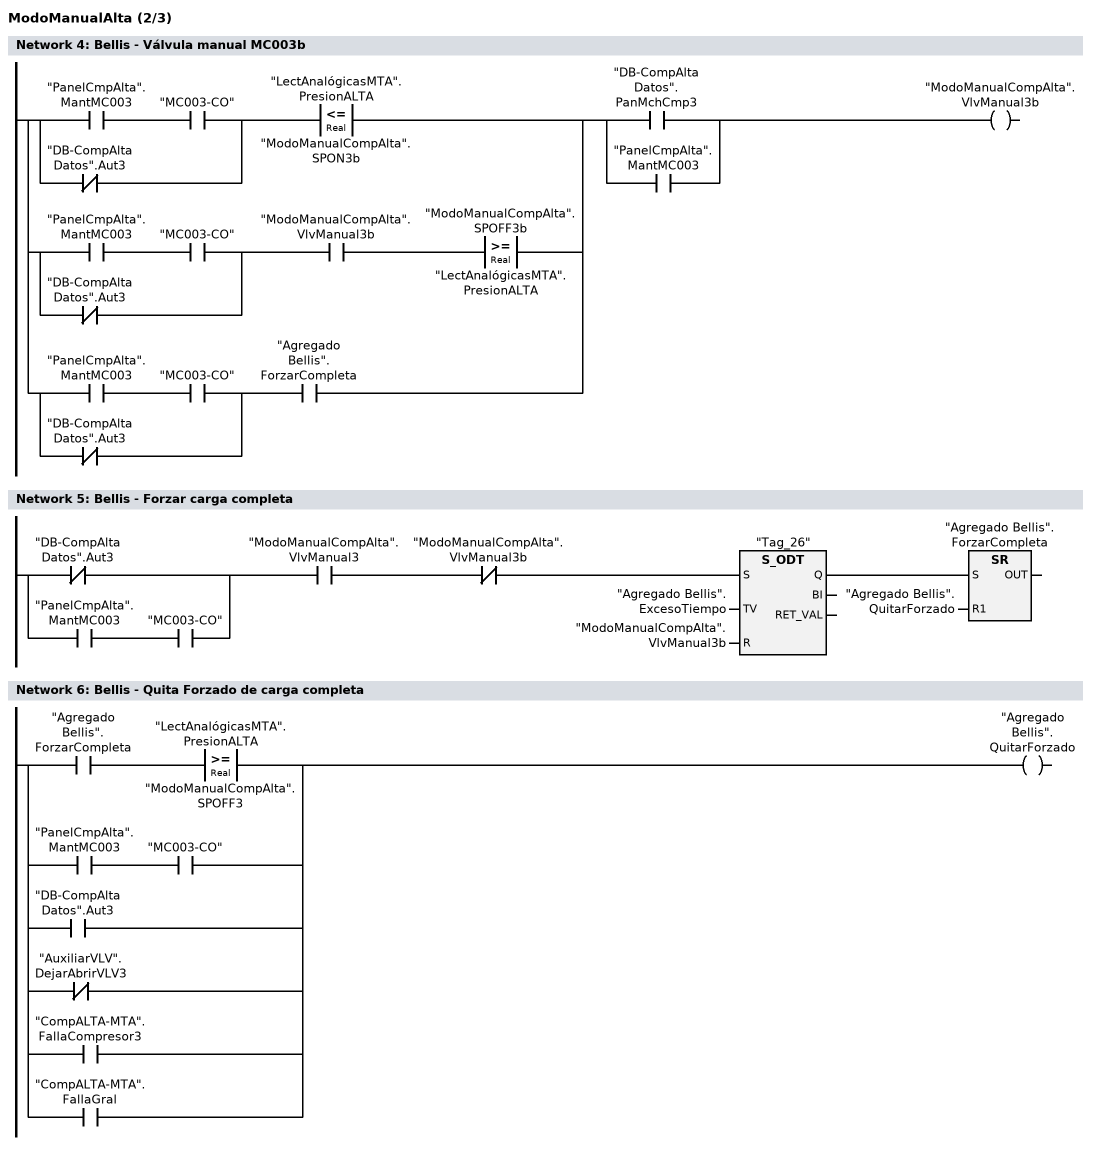
   "ModoManualCompAlta".VlvManual3b := (((NOT "DB-CompAltaDatos".Aut3 OR ("PanelCmpAlta".MantMC003 AND "MC003-CO")) AND ("LectAnalógicasMTA".PresionALTA <= "ModoManualCompAlta".SPON3b)) OR ((NOT "DB-CompAltaDatos".Aut3 OR ("PanelCmpAlta".MantMC003 AND "MC003-CO")) AND "ModoManualCompAlta".VlvManual3b AND ("ModoManualCompAlta".SPOFF3b >= "LectAnalógicasMTA".PresionALTA)) OR ((NOT "DB-CompAltaDatos".Aut3 OR ("PanelCmpAlta".MantMC003 AND "MC003-CO")) AND "Agregado Bellis".ForzarCompleta)) AND ("DB-CompAltaDatos".PanMchCmp3 OR "PanelCmpAlta".MantMC003);
END_REGION

REGION Network 5: Bellis - Forzar carga completa
   RUNG wire#powerrail
      I_Contact( "DB-CompAltaDatos".Aut3 )
      wire#w1
      Contact( "ModoManualCompAlta".VlvManual3 )
      I_Contact( "ModoManualCompAlta".VlvManual3b )
      S_ODT(T_NO := "Tag_26", TV := "Agregado Bellis".ExcesoTiempo, R := "ModoManualCompAlta".VlvManual3b, BI =>, RET_VAL =>)
      S_SR(operand := "Agregado Bellis".ForzarCompleta, r1 := "Agregado Bellis".QuitarForzado)
   END_RUNG
   RUNG wire#powerrail
      Contact( "PanelCmpAlta".MantMC003 )
      Contact( "MC003-CO" )
   END_RUNG wire#w1
   // the same network as SCL:
   #_s5time1 := S_ODT(T_NO := "Tag_26",
                      S := (NOT "DB-CompAltaDatos".Aut3 OR ("PanelCmpAlta".MantMC003 AND "MC003-CO")) AND "ModoManualCompAlta".VlvManual3 AND NOT "ModoManualCompAlta".VlvManual3b,
                      TV := "Agregado Bellis".ExcesoTiempo,
                      R := "ModoManualCompAlta".VlvManual3b,
                      Q => #_w1);
   IF #_w1 THEN
       "Agregado Bellis".ForzarCompleta := TRUE;   // SR flip-flop
   END_IF;
   IF "Agregado Bellis".QuitarForzado THEN "Agregado Bellis".ForzarCompleta := FALSE; END_IF;
END_REGION

REGION Network 6: Bellis - Quita Forzado de carga completa
   "Agregado Bellis".QuitarForzado := ("Agregado Bellis".ForzarCompleta AND ("LectAnalógicasMTA".PresionALTA >= "ModoManualCompAlta".SPOFF3)) OR "DB-CompAltaDatos".Aut3 OR ("PanelCmpAlta".MantMC003 AND "MC003-CO") OR NOT "AuxiliarVLV".DejarAbrirVLV3 OR "CompALTA-MTA".FallaCompresor3 OR "CompALTA-MTA".FallaGral;
END_REGION

REGION Network 7
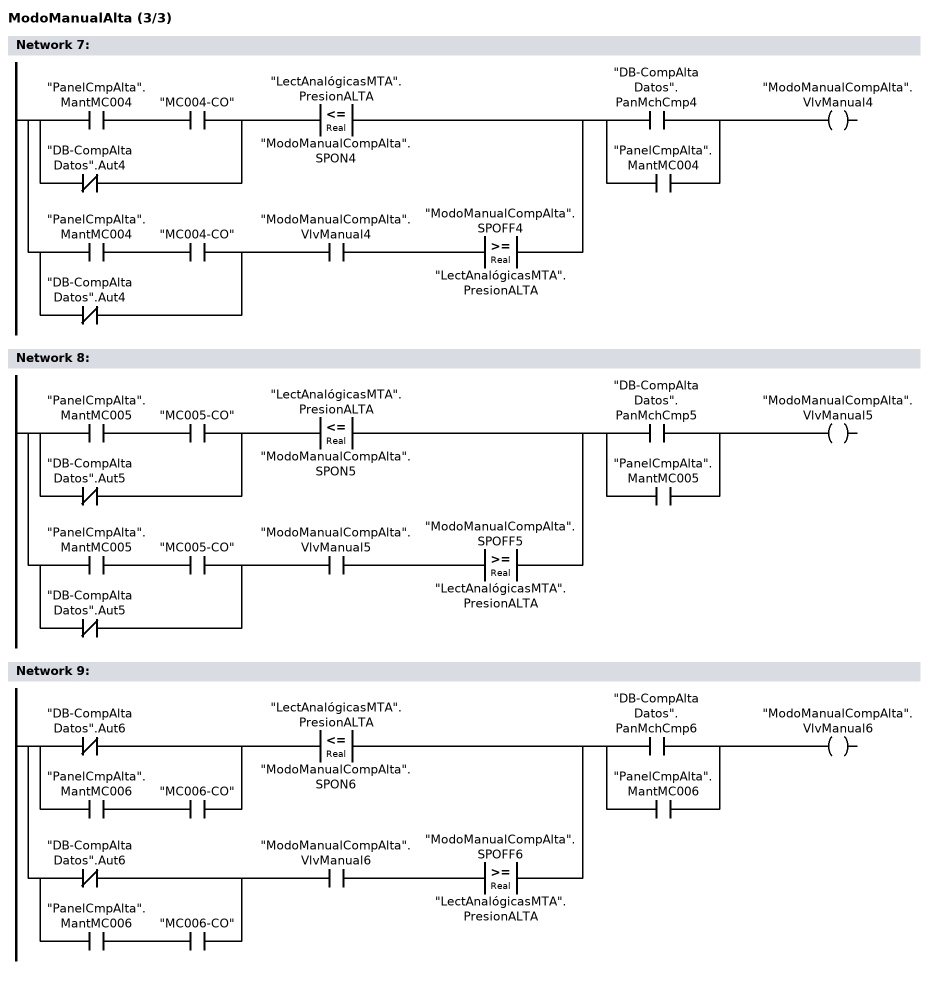
   "ModoManualCompAlta".VlvManual4 := (((NOT "DB-CompAltaDatos".Aut4 OR ("PanelCmpAlta".MantMC004 AND "MC004-CO")) AND ("LectAnalógicasMTA".PresionALTA <= "ModoManualCompAlta".SPON4)) OR ((NOT "DB-CompAltaDatos".Aut4 OR ("PanelCmpAlta".MantMC004 AND "MC004-CO")) AND "ModoManualCompAlta".VlvManual4 AND ("ModoManualCompAlta".SPOFF4 >= "LectAnalógicasMTA".PresionALTA))) AND ("DB-CompAltaDatos".PanMchCmp4 OR "PanelCmpAlta".MantMC004);
END_REGION

REGION Network 8
   "ModoManualCompAlta".VlvManual5 := (((NOT "DB-CompAltaDatos".Aut5 OR ("PanelCmpAlta".MantMC005 AND "MC005-CO")) AND ("LectAnalógicasMTA".PresionALTA <= "ModoManualCompAlta".SPON5)) OR ((NOT "DB-CompAltaDatos".Aut5 OR ("PanelCmpAlta".MantMC005 AND "MC005-CO")) AND "ModoManualCompAlta".VlvManual5 AND ("ModoManualCompAlta".SPOFF5 >= "LectAnalógicasMTA".PresionALTA))) AND ("DB-CompAltaDatos".PanMchCmp5 OR "PanelCmpAlta".MantMC005);
END_REGION

REGION Network 9
   RUNG wire#powerrail
      I_Contact( "DB-CompAltaDatos".Aut6 )
      wire#w1
      { S7_Templates := "SrcType := Real" } LE_Contact(in1 := "LectAnalógicasMTA".PresionALTA, in2 := "ModoManualCompAlta".SPON6)
      wire#w2
      Contact( "DB-CompAltaDatos".PanMchCmp6 )
      wire#w4
      Coil( "ModoManualCompAlta".VlvManual6 )
   END_RUNG
   RUNG wire#powerrail
      Contact( "PanelCmpAlta".MantMC006 )
      Contact( "MC006-CO" )
   END_RUNG wire#w1
   RUNG wire#powerrail
      I_Contact( "DB-CompAltaDatos".Aut6 )
      wire#w3
      Contact( "ModoManualCompAlta".VlvManual6 )
      { S7_Templates := "SrcType := Real" } GE_Contact(in1 := "ModoManualCompAlta".SPOFF6, in2 := "LectAnalógicasMTA".PresionALTA)
   END_RUNG wire#w2
   RUNG wire#powerrail
      Contact( "PanelCmpAlta".MantMC006 )
      Contact( "MC006-CO" )
   END_RUNG wire#w3
   RUNG wire#w2
      Contact( "PanelCmpAlta".MantMC006 )
   END_RUNG wire#w4
   // the same network as SCL:
   "ModoManualCompAlta".VlvManual6 := (((NOT "DB-CompAltaDatos".Aut6 OR ("PanelCmpAlta".MantMC006 AND "MC006-CO")) AND ("LectAnalógicasMTA".PresionALTA <= "ModoManualCompAlta".SPON6)) OR ((NOT "DB-CompAltaDatos".Aut6 OR ("PanelCmpAlta".MantMC006 AND "MC006-CO")) AND "ModoManualCompAlta".VlvManual6 AND ("ModoManualCompAlta".SPOFF6 >= "LectAnalógicasMTA".PresionALTA))) AND ("DB-CompAltaDatos".PanMchCmp6 OR "PanelCmpAlta".MantMC006);
END_REGION
END_FUNCTION

// folder: Compresores/Alta/Máquina de Estados

FUNCTION "LogMaqEstGeneral" : Void   // FC35, LAD
{ S7_Optimized_Access := 'FALSE' }
VERSION : 0.1
BEGIN

REGION Network 1
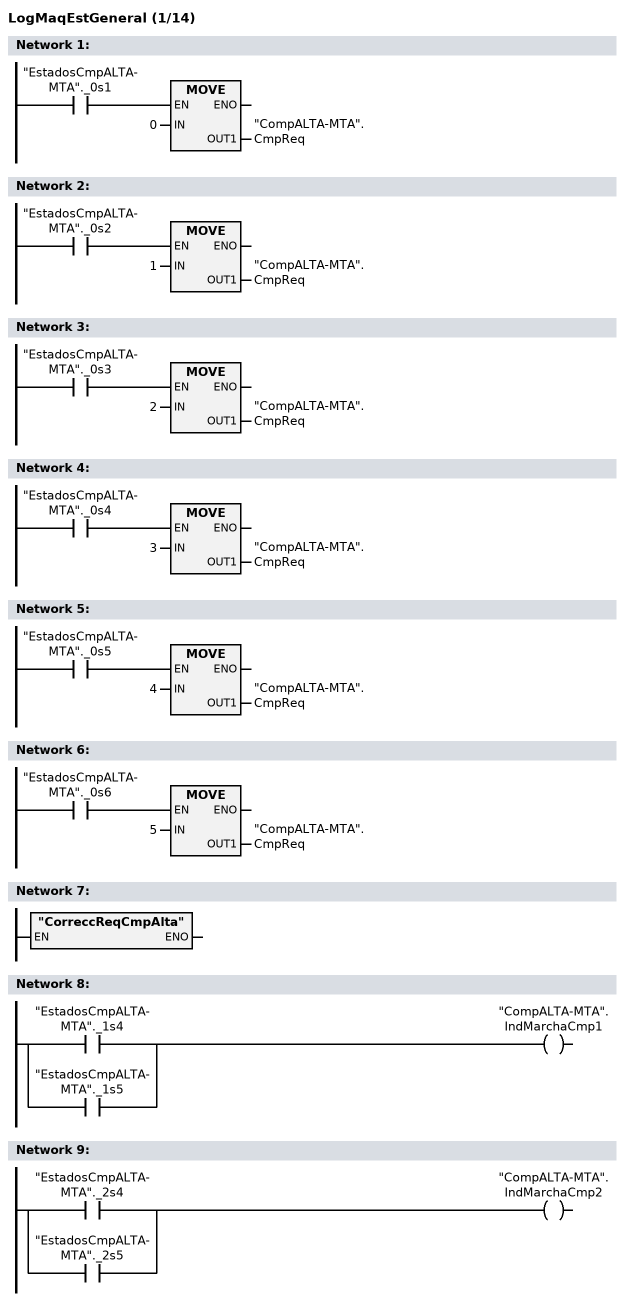
   RUNG wire#powerrail
      Contact( "EstadosCmpALTA-MTA"._0s1 )
      { S7_GenerateENO := "TRUE" } Move(in := 0, out1 => "CompALTA-MTA".CmpReq)
   END_RUNG
   // the same network as SCL:
   IF "EstadosCmpALTA-MTA"._0s1 THEN "CompALTA-MTA".CmpReq := 0; END_IF;
END_REGION

REGION Network 2
   RUNG wire#powerrail
      Contact( "EstadosCmpALTA-MTA"._0s2 )
      { S7_GenerateENO := "TRUE" } Move(in := 1, out1 => "CompALTA-MTA".CmpReq)
   END_RUNG
   // the same network as SCL:
   IF "EstadosCmpALTA-MTA"._0s2 THEN "CompALTA-MTA".CmpReq := 1; END_IF;
END_REGION

REGION Network 3
   RUNG wire#powerrail
      Contact( "EstadosCmpALTA-MTA"._0s3 )
      { S7_GenerateENO := "TRUE" } Move(in := 2, out1 => "CompALTA-MTA".CmpReq)
   END_RUNG
   // the same network as SCL:
   IF "EstadosCmpALTA-MTA"._0s3 THEN "CompALTA-MTA".CmpReq := 2; END_IF;
END_REGION

REGION Network 4
   RUNG wire#powerrail
      Contact( "EstadosCmpALTA-MTA"._0s4 )
      { S7_GenerateENO := "TRUE" } Move(in := 3, out1 => "CompALTA-MTA".CmpReq)
   END_RUNG
   // the same network as SCL:
   IF "EstadosCmpALTA-MTA"._0s4 THEN "CompALTA-MTA".CmpReq := 3; END_IF;
END_REGION

REGION Network 5
   RUNG wire#powerrail
      Contact( "EstadosCmpALTA-MTA"._0s5 )
      { S7_GenerateENO := "TRUE" } Move(in := 4, out1 => "CompALTA-MTA".CmpReq)
   END_RUNG
   // the same network as SCL:
   IF "EstadosCmpALTA-MTA"._0s5 THEN "CompALTA-MTA".CmpReq := 4; END_IF;
END_REGION

REGION Network 6
   RUNG wire#powerrail
      Contact( "EstadosCmpALTA-MTA"._0s6 )
      { S7_GenerateENO := "TRUE" } Move(in := 5, out1 => "CompALTA-MTA".CmpReq)
   END_RUNG
   // the same network as SCL:
   IF "EstadosCmpALTA-MTA"._0s6 THEN "CompALTA-MTA".CmpReq := 5; END_IF;
END_REGION

REGION Network 7
   RUNG wire#powerrail
      "CorreccReqCmpAlta"()
   END_RUNG
   // the same network as SCL:
   "CorreccReqCmpAlta"();
END_REGION

REGION Network 8
   RUNG wire#powerrail
      Contact( "EstadosCmpALTA-MTA"._1s4 )
      wire#w1
      Coil( "CompALTA-MTA".IndMarchaCmp1 )
   END_RUNG
   RUNG wire#powerrail
      Contact( "EstadosCmpALTA-MTA"._1s5 )
   END_RUNG wire#w1
   // the same network as SCL:
   "CompALTA-MTA".IndMarchaCmp1 := "EstadosCmpALTA-MTA"._1s4 OR "EstadosCmpALTA-MTA"._1s5;
END_REGION

REGION Network 9
   RUNG wire#powerrail
      Contact( "EstadosCmpALTA-MTA"._2s4 )
      wire#w1
      Coil( "CompALTA-MTA".IndMarchaCmp2 )
   END_RUNG
   RUNG wire#powerrail
      Contact( "EstadosCmpALTA-MTA"._2s5 )
   END_RUNG wire#w1
   // the same network as SCL:
   "CompALTA-MTA".IndMarchaCmp2 := "EstadosCmpALTA-MTA"._2s4 OR "EstadosCmpALTA-MTA"._2s5;
END_REGION

REGION Network 10
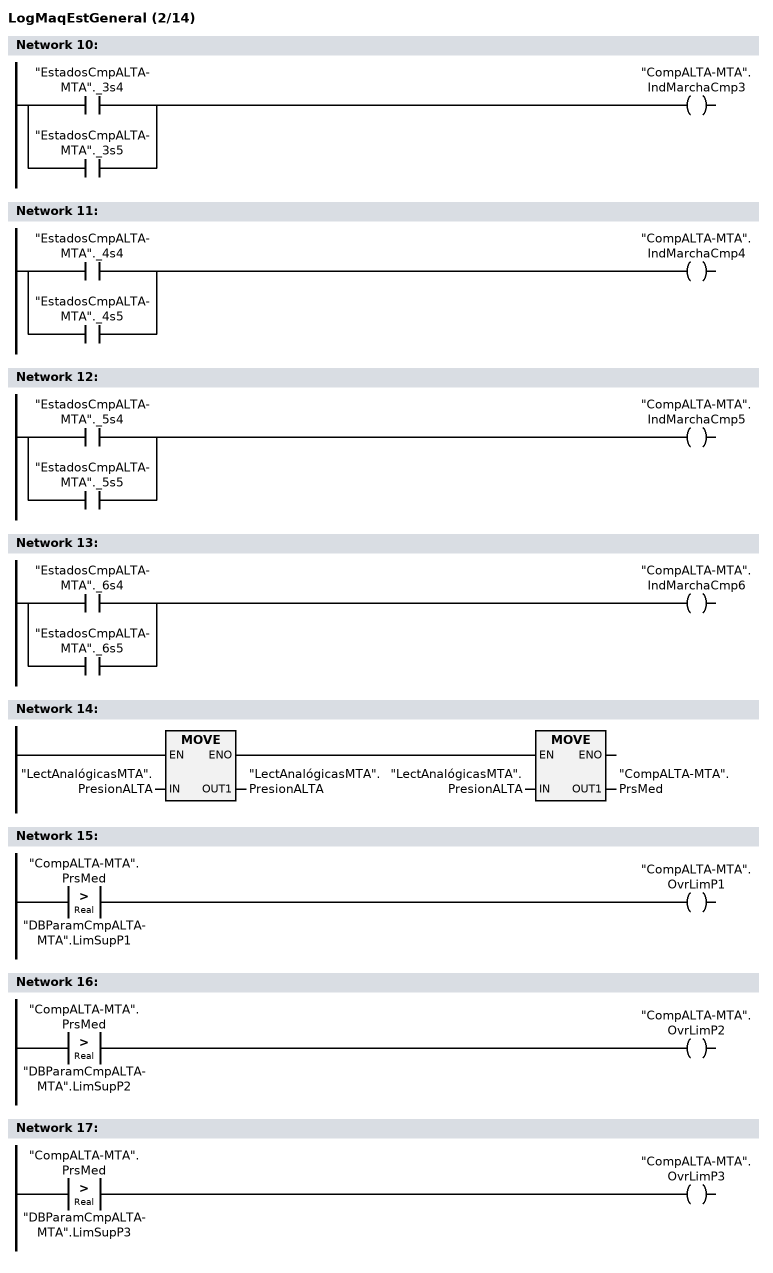
   RUNG wire#powerrail
      Contact( "EstadosCmpALTA-MTA"._3s4 )
      wire#w1
      Coil( "CompALTA-MTA".IndMarchaCmp3 )
   END_RUNG
   RUNG wire#powerrail
      Contact( "EstadosCmpALTA-MTA"._3s5 )
   END_RUNG wire#w1
   // the same network as SCL:
   "CompALTA-MTA".IndMarchaCmp3 := "EstadosCmpALTA-MTA"._3s4 OR "EstadosCmpALTA-MTA"._3s5;
END_REGION

REGION Network 11
   RUNG wire#powerrail
      Contact( "EstadosCmpALTA-MTA"._4s4 )
      wire#w1
      Coil( "CompALTA-MTA".IndMarchaCmp4 )
   END_RUNG
   RUNG wire#powerrail
      Contact( "EstadosCmpALTA-MTA"._4s5 )
   END_RUNG wire#w1
   // the same network as SCL:
   "CompALTA-MTA".IndMarchaCmp4 := "EstadosCmpALTA-MTA"._4s4 OR "EstadosCmpALTA-MTA"._4s5;
END_REGION

REGION Network 12
   RUNG wire#powerrail
      Contact( "EstadosCmpALTA-MTA"._5s4 )
      wire#w1
      Coil( "CompALTA-MTA".IndMarchaCmp5 )
   END_RUNG
   RUNG wire#powerrail
      Contact( "EstadosCmpALTA-MTA"._5s5 )
   END_RUNG wire#w1
   // the same network as SCL:
   "CompALTA-MTA".IndMarchaCmp5 := "EstadosCmpALTA-MTA"._5s4 OR "EstadosCmpALTA-MTA"._5s5;
END_REGION

REGION Network 13
   RUNG wire#powerrail
      Contact( "EstadosCmpALTA-MTA"._6s4 )
      wire#w1
      Coil( "CompALTA-MTA".IndMarchaCmp6 )
   END_RUNG
   RUNG wire#powerrail
      Contact( "EstadosCmpALTA-MTA"._6s5 )
   END_RUNG wire#w1
   // the same network as SCL:
   "CompALTA-MTA".IndMarchaCmp6 := "EstadosCmpALTA-MTA"._6s4 OR "EstadosCmpALTA-MTA"._6s5;
END_REGION

REGION Network 14
   RUNG wire#powerrail
      { S7_GenerateENO := "TRUE" } Move(in := "LectAnalógicasMTA".PresionALTA, out1 => "LectAnalógicasMTA".PresionALTA)
      { S7_GenerateENO := "TRUE" } Move(in := "LectAnalógicasMTA".PresionALTA, out1 => "CompALTA-MTA".PrsMed)
   END_RUNG
   // the same network as SCL:
   // ENO of a box is taken as its EN; it also drops when the box reports an error
   "LectAnalógicasMTA".PresionALTA := "LectAnalógicasMTA".PresionALTA;
   "CompALTA-MTA".PrsMed := "LectAnalógicasMTA".PresionALTA;
END_REGION

REGION Network 15
   RUNG wire#powerrail
      { S7_Templates := "SrcType := Real" } GT_Contact(in1 := "CompALTA-MTA".PrsMed, in2 := "DBParamCmpALTA-MTA".LimSupP1)
      Coil( "CompALTA-MTA".OvrLimP1 )
   END_RUNG
   // the same network as SCL:
   "CompALTA-MTA".OvrLimP1 := "CompALTA-MTA".PrsMed > "DBParamCmpALTA-MTA".LimSupP1;
END_REGION

REGION Network 16
   RUNG wire#powerrail
      { S7_Templates := "SrcType := Real" } GT_Contact(in1 := "CompALTA-MTA".PrsMed, in2 := "DBParamCmpALTA-MTA".LimSupP2)
      Coil( "CompALTA-MTA".OvrLimP2 )
   END_RUNG
   // the same network as SCL:
   "CompALTA-MTA".OvrLimP2 := "CompALTA-MTA".PrsMed > "DBParamCmpALTA-MTA".LimSupP2;
END_REGION

REGION Network 17
   RUNG wire#powerrail
      { S7_Templates := "SrcType := Real" } GT_Contact(in1 := "CompALTA-MTA".PrsMed, in2 := "DBParamCmpALTA-MTA".LimSupP3)
      Coil( "CompALTA-MTA".OvrLimP3 )
   END_RUNG
   // the same network as SCL:
   "CompALTA-MTA".OvrLimP3 := "CompALTA-MTA".PrsMed > "DBParamCmpALTA-MTA".LimSupP3;
END_REGION

REGION Network 18
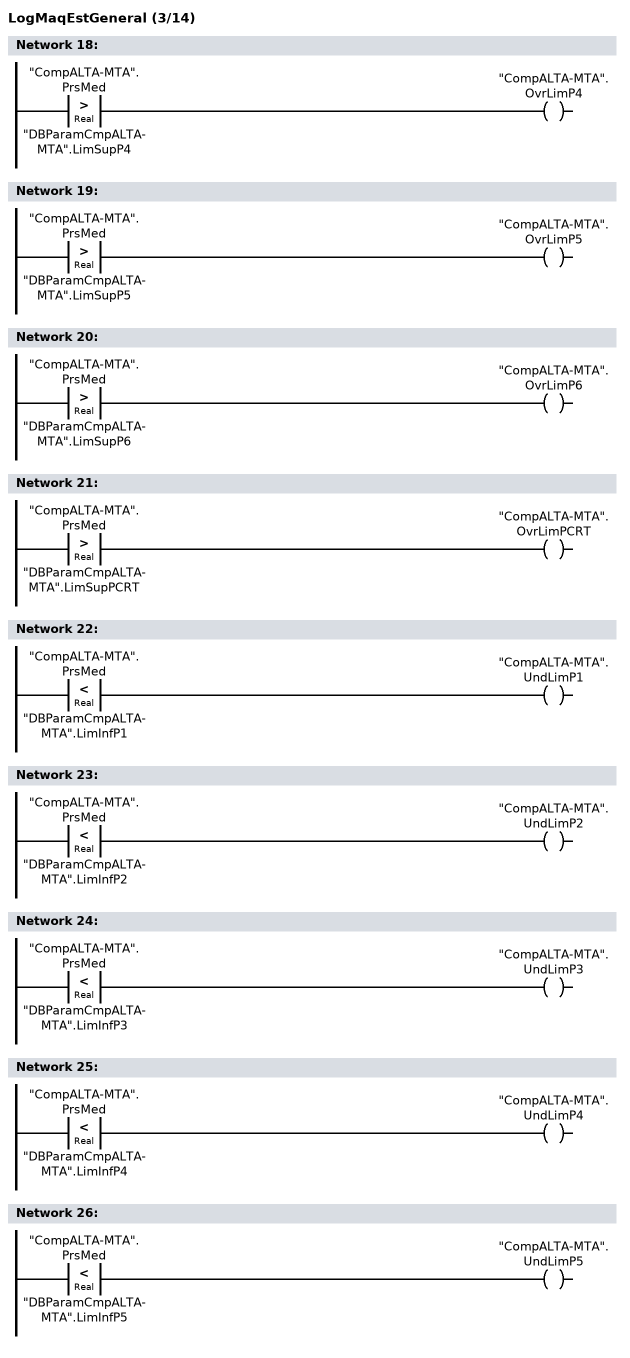
   RUNG wire#powerrail
      { S7_Templates := "SrcType := Real" } GT_Contact(in1 := "CompALTA-MTA".PrsMed, in2 := "DBParamCmpALTA-MTA".LimSupP4)
      Coil( "CompALTA-MTA".OvrLimP4 )
   END_RUNG
   // the same network as SCL:
   "CompALTA-MTA".OvrLimP4 := "CompALTA-MTA".PrsMed > "DBParamCmpALTA-MTA".LimSupP4;
END_REGION

REGION Network 19
   RUNG wire#powerrail
      { S7_Templates := "SrcType := Real" } GT_Contact(in1 := "CompALTA-MTA".PrsMed, in2 := "DBParamCmpALTA-MTA".LimSupP5)
      Coil( "CompALTA-MTA".OvrLimP5 )
   END_RUNG
   // the same network as SCL:
   "CompALTA-MTA".OvrLimP5 := "CompALTA-MTA".PrsMed > "DBParamCmpALTA-MTA".LimSupP5;
END_REGION

REGION Network 20
   RUNG wire#powerrail
      { S7_Templates := "SrcType := Real" } GT_Contact(in1 := "CompALTA-MTA".PrsMed, in2 := "DBParamCmpALTA-MTA".LimSupP6)
      Coil( "CompALTA-MTA".OvrLimP6 )
   END_RUNG
   // the same network as SCL:
   "CompALTA-MTA".OvrLimP6 := "CompALTA-MTA".PrsMed > "DBParamCmpALTA-MTA".LimSupP6;
END_REGION

REGION Network 21
   RUNG wire#powerrail
      { S7_Templates := "SrcType := Real" } GT_Contact(in1 := "CompALTA-MTA".PrsMed, in2 := "DBParamCmpALTA-MTA".LimSupPCRT)
      Coil( "CompALTA-MTA".OvrLimPCRT )
   END_RUNG
   // the same network as SCL:
   "CompALTA-MTA".OvrLimPCRT := "CompALTA-MTA".PrsMed > "DBParamCmpALTA-MTA".LimSupPCRT;
END_REGION

REGION Network 22
   RUNG wire#powerrail
      { S7_Templates := "SrcType := Real" } LT_Contact(in1 := "CompALTA-MTA".PrsMed, in2 := "DBParamCmpALTA-MTA".LimInfP1)
      Coil( "CompALTA-MTA".UndLimP1 )
   END_RUNG
   // the same network as SCL:
   "CompALTA-MTA".UndLimP1 := "CompALTA-MTA".PrsMed < "DBParamCmpALTA-MTA".LimInfP1;
END_REGION

REGION Network 23
   RUNG wire#powerrail
      { S7_Templates := "SrcType := Real" } LT_Contact(in1 := "CompALTA-MTA".PrsMed, in2 := "DBParamCmpALTA-MTA".LimInfP2)
      Coil( "CompALTA-MTA".UndLimP2 )
   END_RUNG
   // the same network as SCL:
   "CompALTA-MTA".UndLimP2 := "CompALTA-MTA".PrsMed < "DBParamCmpALTA-MTA".LimInfP2;
END_REGION

REGION Network 24
   RUNG wire#powerrail
      { S7_Templates := "SrcType := Real" } LT_Contact(in1 := "CompALTA-MTA".PrsMed, in2 := "DBParamCmpALTA-MTA".LimInfP3)
      Coil( "CompALTA-MTA".UndLimP3 )
   END_RUNG
   // the same network as SCL:
   "CompALTA-MTA".UndLimP3 := "CompALTA-MTA".PrsMed < "DBParamCmpALTA-MTA".LimInfP3;
END_REGION

REGION Network 25
   RUNG wire#powerrail
      { S7_Templates := "SrcType := Real" } LT_Contact(in1 := "CompALTA-MTA".PrsMed, in2 := "DBParamCmpALTA-MTA".LimInfP4)
      Coil( "CompALTA-MTA".UndLimP4 )
   END_RUNG
   // the same network as SCL:
   "CompALTA-MTA".UndLimP4 := "CompALTA-MTA".PrsMed < "DBParamCmpALTA-MTA".LimInfP4;
END_REGION

REGION Network 26
   RUNG wire#powerrail
      { S7_Templates := "SrcType := Real" } LT_Contact(in1 := "CompALTA-MTA".PrsMed, in2 := "DBParamCmpALTA-MTA".LimInfP5)
      Coil( "CompALTA-MTA".UndLimP5 )
   END_RUNG
   // the same network as SCL:
   "CompALTA-MTA".UndLimP5 := "CompALTA-MTA".PrsMed < "DBParamCmpALTA-MTA".LimInfP5;
END_REGION

REGION Network 27
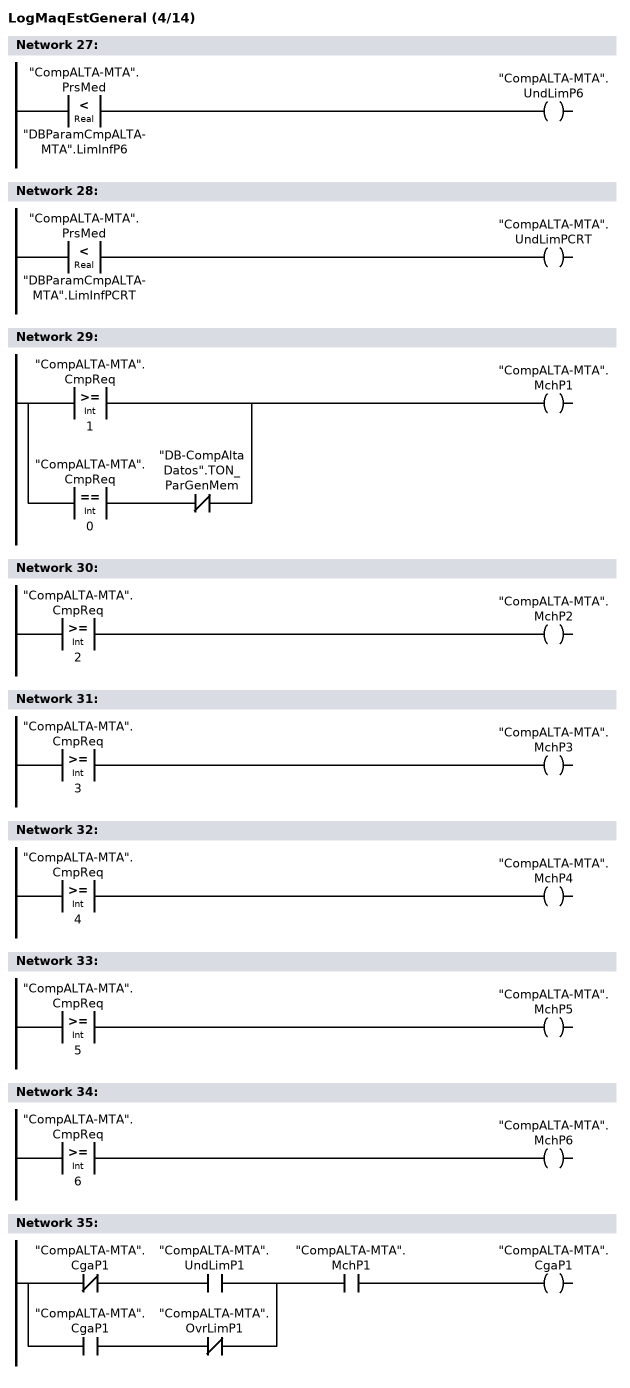
   RUNG wire#powerrail
      { S7_Templates := "SrcType := Real" } LT_Contact(in1 := "CompALTA-MTA".PrsMed, in2 := "DBParamCmpALTA-MTA".LimInfP6)
      Coil( "CompALTA-MTA".UndLimP6 )
   END_RUNG
   // the same network as SCL:
   "CompALTA-MTA".UndLimP6 := "CompALTA-MTA".PrsMed < "DBParamCmpALTA-MTA".LimInfP6;
END_REGION

REGION Network 28
   RUNG wire#powerrail
      { S7_Templates := "SrcType := Real" } LT_Contact(in1 := "CompALTA-MTA".PrsMed, in2 := "DBParamCmpALTA-MTA".LimInfPCRT)
      Coil( "CompALTA-MTA".UndLimPCRT )
   END_RUNG
   // the same network as SCL:
   "CompALTA-MTA".UndLimPCRT := "CompALTA-MTA".PrsMed < "DBParamCmpALTA-MTA".LimInfPCRT;
END_REGION

REGION Network 29
   RUNG wire#powerrail
      { S7_Templates := "SrcType := Int" } GE_Contact(in1 := "CompALTA-MTA".CmpReq, in2 := 1)
      wire#w1
      Coil( "CompALTA-MTA".MchP1 )
   END_RUNG
   RUNG wire#powerrail
      { S7_Templates := "SrcType := Int" } EQ_Contact(in1 := "CompALTA-MTA".CmpReq, in2 := 0)
      I_Contact( "DB-CompAltaDatos".TON_ParGenMem )
   END_RUNG wire#w1
   // the same network as SCL:
   "CompALTA-MTA".MchP1 := ("CompALTA-MTA".CmpReq >= 1) OR (("CompALTA-MTA".CmpReq = 0) AND NOT "DB-CompAltaDatos".TON_ParGenMem);
END_REGION

REGION Network 30
   RUNG wire#powerrail
      { S7_Templates := "SrcType := Int" } GE_Contact(in1 := "CompALTA-MTA".CmpReq, in2 := 2)
      Coil( "CompALTA-MTA".MchP2 )
   END_RUNG
   // the same network as SCL:
   "CompALTA-MTA".MchP2 := "CompALTA-MTA".CmpReq >= 2;
END_REGION

REGION Network 31
   RUNG wire#powerrail
      { S7_Templates := "SrcType := Int" } GE_Contact(in1 := "CompALTA-MTA".CmpReq, in2 := 3)
      Coil( "CompALTA-MTA".MchP3 )
   END_RUNG
   // the same network as SCL:
   "CompALTA-MTA".MchP3 := "CompALTA-MTA".CmpReq >= 3;
END_REGION

REGION Network 32
   RUNG wire#powerrail
      { S7_Templates := "SrcType := Int" } GE_Contact(in1 := "CompALTA-MTA".CmpReq, in2 := 4)
      Coil( "CompALTA-MTA".MchP4 )
   END_RUNG
   // the same network as SCL:
   "CompALTA-MTA".MchP4 := "CompALTA-MTA".CmpReq >= 4;
END_REGION

REGION Network 33
   RUNG wire#powerrail
      { S7_Templates := "SrcType := Int" } GE_Contact(in1 := "CompALTA-MTA".CmpReq, in2 := 5)
      Coil( "CompALTA-MTA".MchP5 )
   END_RUNG
   // the same network as SCL:
   "CompALTA-MTA".MchP5 := "CompALTA-MTA".CmpReq >= 5;
END_REGION

REGION Network 34
   RUNG wire#powerrail
      { S7_Templates := "SrcType := Int" } GE_Contact(in1 := "CompALTA-MTA".CmpReq, in2 := 6)
      Coil( "CompALTA-MTA".MchP6 )
   END_RUNG
   // the same network as SCL:
   "CompALTA-MTA".MchP6 := "CompALTA-MTA".CmpReq >= 6;
END_REGION

REGION Network 35
   RUNG wire#powerrail
      I_Contact( "CompALTA-MTA".CgaP1 )
      Contact( "CompALTA-MTA".UndLimP1 )
      wire#w1
      Contact( "CompALTA-MTA".MchP1 )
      Coil( "CompALTA-MTA".CgaP1 )
   END_RUNG
   RUNG wire#powerrail
      Contact( "CompALTA-MTA".CgaP1 )
      I_Contact( "CompALTA-MTA".OvrLimP1 )
   END_RUNG wire#w1
   // the same network as SCL:
   "CompALTA-MTA".CgaP1 := ((NOT "CompALTA-MTA".CgaP1 AND "CompALTA-MTA".UndLimP1) OR ("CompALTA-MTA".CgaP1 AND NOT "CompALTA-MTA".OvrLimP1)) AND "CompALTA-MTA".MchP1;
END_REGION

REGION Network 36
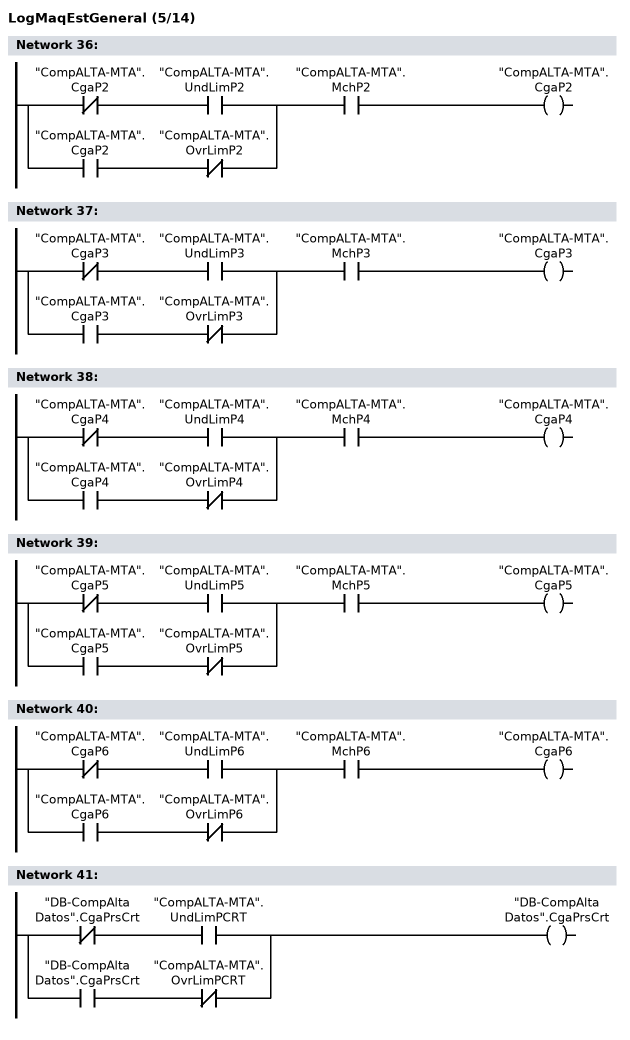
   RUNG wire#powerrail
      I_Contact( "CompALTA-MTA".CgaP2 )
      Contact( "CompALTA-MTA".UndLimP2 )
      wire#w1
      Contact( "CompALTA-MTA".MchP2 )
      Coil( "CompALTA-MTA".CgaP2 )
   END_RUNG
   RUNG wire#powerrail
      Contact( "CompALTA-MTA".CgaP2 )
      I_Contact( "CompALTA-MTA".OvrLimP2 )
   END_RUNG wire#w1
   // the same network as SCL:
   "CompALTA-MTA".CgaP2 := ((NOT "CompALTA-MTA".CgaP2 AND "CompALTA-MTA".UndLimP2) OR ("CompALTA-MTA".CgaP2 AND NOT "CompALTA-MTA".OvrLimP2)) AND "CompALTA-MTA".MchP2;
END_REGION

REGION Network 37
   RUNG wire#powerrail
      I_Contact( "CompALTA-MTA".CgaP3 )
      Contact( "CompALTA-MTA".UndLimP3 )
      wire#w1
      Contact( "CompALTA-MTA".MchP3 )
      Coil( "CompALTA-MTA".CgaP3 )
   END_RUNG
   RUNG wire#powerrail
      Contact( "CompALTA-MTA".CgaP3 )
      I_Contact( "CompALTA-MTA".OvrLimP3 )
   END_RUNG wire#w1
   // the same network as SCL:
   "CompALTA-MTA".CgaP3 := ((NOT "CompALTA-MTA".CgaP3 AND "CompALTA-MTA".UndLimP3) OR ("CompALTA-MTA".CgaP3 AND NOT "CompALTA-MTA".OvrLimP3)) AND "CompALTA-MTA".MchP3;
END_REGION

REGION Network 38
   RUNG wire#powerrail
      I_Contact( "CompALTA-MTA".CgaP4 )
      Contact( "CompALTA-MTA".UndLimP4 )
      wire#w1
      Contact( "CompALTA-MTA".MchP4 )
      Coil( "CompALTA-MTA".CgaP4 )
   END_RUNG
   RUNG wire#powerrail
      Contact( "CompALTA-MTA".CgaP4 )
      I_Contact( "CompALTA-MTA".OvrLimP4 )
   END_RUNG wire#w1
   // the same network as SCL:
   "CompALTA-MTA".CgaP4 := ((NOT "CompALTA-MTA".CgaP4 AND "CompALTA-MTA".UndLimP4) OR ("CompALTA-MTA".CgaP4 AND NOT "CompALTA-MTA".OvrLimP4)) AND "CompALTA-MTA".MchP4;
END_REGION

REGION Network 39
   RUNG wire#powerrail
      I_Contact( "CompALTA-MTA".CgaP5 )
      Contact( "CompALTA-MTA".UndLimP5 )
      wire#w1
      Contact( "CompALTA-MTA".MchP5 )
      Coil( "CompALTA-MTA".CgaP5 )
   END_RUNG
   RUNG wire#powerrail
      Contact( "CompALTA-MTA".CgaP5 )
      I_Contact( "CompALTA-MTA".OvrLimP5 )
   END_RUNG wire#w1
   // the same network as SCL:
   "CompALTA-MTA".CgaP5 := ((NOT "CompALTA-MTA".CgaP5 AND "CompALTA-MTA".UndLimP5) OR ("CompALTA-MTA".CgaP5 AND NOT "CompALTA-MTA".OvrLimP5)) AND "CompALTA-MTA".MchP5;
END_REGION

REGION Network 40
   RUNG wire#powerrail
      I_Contact( "CompALTA-MTA".CgaP6 )
      Contact( "CompALTA-MTA".UndLimP6 )
      wire#w1
      Contact( "CompALTA-MTA".MchP6 )
      Coil( "CompALTA-MTA".CgaP6 )
   END_RUNG
   RUNG wire#powerrail
      Contact( "CompALTA-MTA".CgaP6 )
      I_Contact( "CompALTA-MTA".OvrLimP6 )
   END_RUNG wire#w1
   // the same network as SCL:
   "CompALTA-MTA".CgaP6 := ((NOT "CompALTA-MTA".CgaP6 AND "CompALTA-MTA".UndLimP6) OR ("CompALTA-MTA".CgaP6 AND NOT "CompALTA-MTA".OvrLimP6)) AND "CompALTA-MTA".MchP6;
END_REGION

REGION Network 41
   RUNG wire#powerrail
      I_Contact( "DB-CompAltaDatos".CgaPrsCrt )
      Contact( "CompALTA-MTA".UndLimPCRT )
      wire#w1
      Coil( "DB-CompAltaDatos".CgaPrsCrt )
   END_RUNG
   RUNG wire#powerrail
      Contact( "DB-CompAltaDatos".CgaPrsCrt )
      I_Contact( "CompALTA-MTA".OvrLimPCRT )
   END_RUNG wire#w1
   // the same network as SCL:
   "DB-CompAltaDatos".CgaPrsCrt := (NOT "DB-CompAltaDatos".CgaPrsCrt AND "CompALTA-MTA".UndLimPCRT) OR ("DB-CompAltaDatos".CgaPrsCrt AND NOT "CompALTA-MTA".OvrLimPCRT);
END_REGION

REGION Network 42
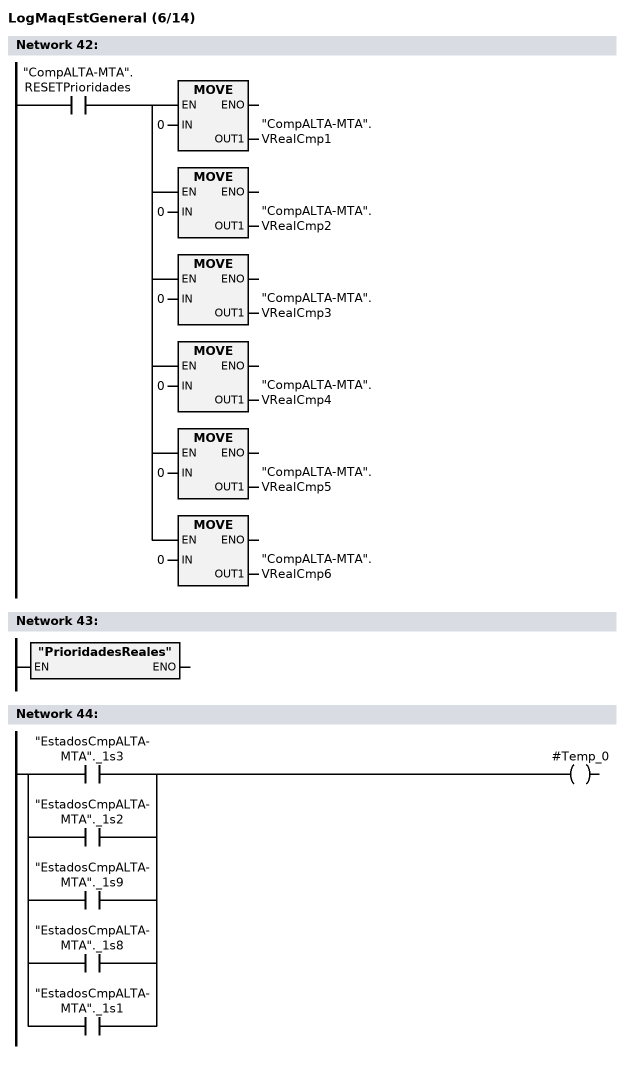
   RUNG wire#powerrail
      Contact( "CompALTA-MTA".RESETPrioridades )
      wire#w1
      { S7_GenerateENO := "TRUE" } Move(in := 0, out1 => "CompALTA-MTA".VRealCmp1)
   END_RUNG
   RUNG wire#w1
      { S7_GenerateENO := "TRUE" } Move(in := 0, out1 => "CompALTA-MTA".VRealCmp2)
   END_RUNG
   RUNG wire#w1
      { S7_GenerateENO := "TRUE" } Move(in := 0, out1 => "CompALTA-MTA".VRealCmp3)
   END_RUNG
   RUNG wire#w1
      { S7_GenerateENO := "TRUE" } Move(in := 0, out1 => "CompALTA-MTA".VRealCmp4)
   END_RUNG
   RUNG wire#w1
      { S7_GenerateENO := "TRUE" } Move(in := 0, out1 => "CompALTA-MTA".VRealCmp5)
   END_RUNG
   RUNG wire#w1
      { S7_GenerateENO := "TRUE" } Move(in := 0, out1 => "CompALTA-MTA".VRealCmp6)
   END_RUNG
   // the same network as SCL:
   IF "CompALTA-MTA".RESETPrioridades THEN
       "CompALTA-MTA".VRealCmp1 := 0;
       "CompALTA-MTA".VRealCmp2 := 0;
       "CompALTA-MTA".VRealCmp3 := 0;
       "CompALTA-MTA".VRealCmp4 := 0;
       "CompALTA-MTA".VRealCmp5 := 0;
       "CompALTA-MTA".VRealCmp6 := 0;
   END_IF;
END_REGION

REGION Network 43
   RUNG wire#powerrail
      "PrioridadesReales"()
   END_RUNG
   // the same network as SCL:
   "PrioridadesReales"();
END_REGION

REGION Network 44
   RUNG wire#powerrail
      Contact( "EstadosCmpALTA-MTA"._1s3 )
      wire#w1
      Coil( #Temp_0 )
   END_RUNG
   RUNG wire#powerrail
      Contact( "EstadosCmpALTA-MTA"._1s2 )
   END_RUNG wire#w1
   RUNG wire#powerrail
      Contact( "EstadosCmpALTA-MTA"._1s9 )
   END_RUNG wire#w1
   RUNG wire#powerrail
      Contact( "EstadosCmpALTA-MTA"._1s8 )
   END_RUNG wire#w1
   RUNG wire#powerrail
      Contact( "EstadosCmpALTA-MTA"._1s1 )
   END_RUNG wire#w1
   // the same network as SCL:
   #Temp_0 := "EstadosCmpALTA-MTA"._1s3 OR "EstadosCmpALTA-MTA"._1s2 OR "EstadosCmpALTA-MTA"._1s9 OR "EstadosCmpALTA-MTA"._1s8 OR "EstadosCmpALTA-MTA"._1s1;
END_REGION

REGION Network 45
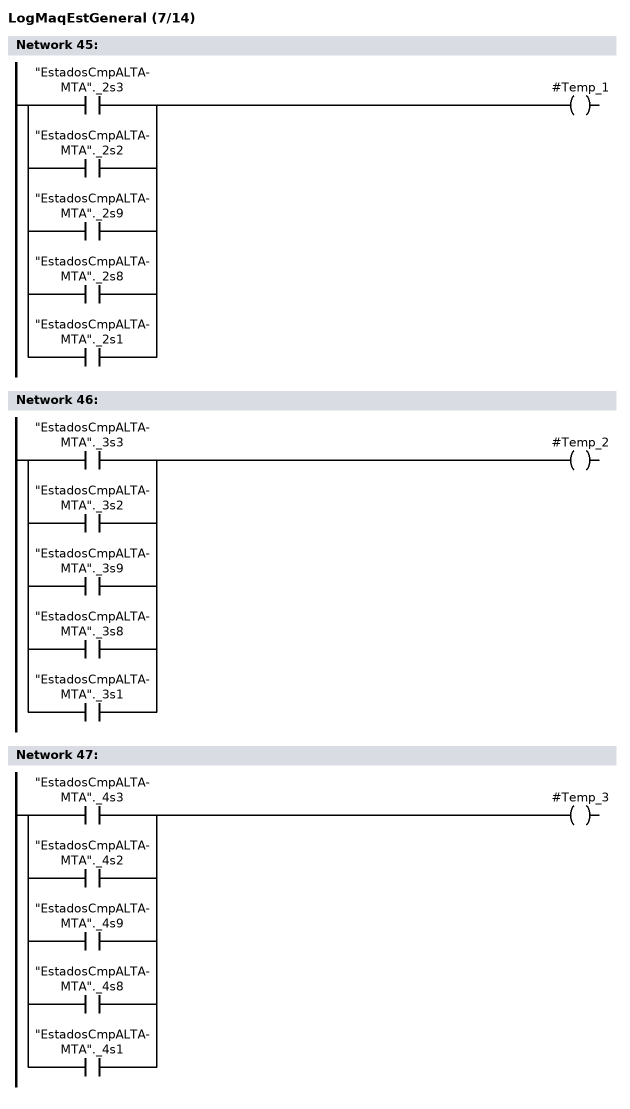
   RUNG wire#powerrail
      Contact( "EstadosCmpALTA-MTA"._2s3 )
      wire#w1
      Coil( #Temp_1 )
   END_RUNG
   RUNG wire#powerrail
      Contact( "EstadosCmpALTA-MTA"._2s2 )
   END_RUNG wire#w1
   RUNG wire#powerrail
      Contact( "EstadosCmpALTA-MTA"._2s9 )
   END_RUNG wire#w1
   RUNG wire#powerrail
      Contact( "EstadosCmpALTA-MTA"._2s8 )
   END_RUNG wire#w1
   RUNG wire#powerrail
      Contact( "EstadosCmpALTA-MTA"._2s1 )
   END_RUNG wire#w1
   // the same network as SCL:
   #Temp_1 := "EstadosCmpALTA-MTA"._2s3 OR "EstadosCmpALTA-MTA"._2s2 OR "EstadosCmpALTA-MTA"._2s9 OR "EstadosCmpALTA-MTA"._2s8 OR "EstadosCmpALTA-MTA"._2s1;
END_REGION
